REGION Network 10: Main Water Pump
   RUNG wire#powerrail
      #VFD_WaterPump(tInTimeout := t#5s, iInMode := #iInMode, iInAddress := 100, bInEstop := #bInEstop, bInSignalContactor := "I_WaterPumpContactorAux", bInEnableForward := #bWaterPumpInterlockOk, bInEnableReverse := false, rInCommandSpeed := 80.0, rInRampUpTime := 5.0, rInRampDownTime := 5.0, bInCommandForward := #bStartPumpCommand, bInCommandReverse := false, bInResetError := #bInResetError, bInMotorProtector := "I_WaterPumpMSP", bInLocalDisconnect := "I_WaterPumpDisconnect", bInClutch := true, bInCoolingFan := "I_WaterPumpCoolingFan", bInUseCurrentAlarm := true, bInUseMaxFrequencyAlarm := true, HMI_VFD_Control := "dbWaterSystem".VFD_WaterPump, rOutSpeed => #rPumpActualSpeed, rOutCurrent => #rPumpActualCurrent, rOutPower => #rPumpActualPower, bOutContactor => "Q_WaterPumpContactor", bOutForward => #bTemp, bOutReverse => #bTemp, bOutAuto => #bTemp, bOutError => #bTemp, ERROR_VFD => "dbErrors_WaterSystem".VFD_WaterPump)
   END_RUNG
   // the same network as SCL:
   #VFD_WaterPump(tInTimeout := t#5s,   // "fbVFD_GSeries"
                  iInMode := #iInMode,
                  iInAddress := 100,
                  bInEstop := #bInEstop,
                  bInSignalContactor := "I_WaterPumpContactorAux",
                  bInEnableForward := #bWaterPumpInterlockOk,
                  bInEnableReverse := false,
                  rInCommandSpeed := 80.0,
                  rInRampUpTime := 5.0,
                  rInRampDownTime := 5.0,
                  bInCommandForward := #bStartPumpCommand,
                  bInCommandReverse := false,
                  bInResetError := #bInResetError,
                  bInMotorProtector := "I_WaterPumpMSP",
                  bInLocalDisconnect := "I_WaterPumpDisconnect",
                  bInClutch := true,
                  bInCoolingFan := "I_WaterPumpCoolingFan",
                  bInUseCurrentAlarm := true,
                  bInUseMaxFrequencyAlarm := true,
                  HMI_VFD_Control := "dbWaterSystem".VFD_WaterPump,
                  rOutSpeed => #rPumpActualSpeed,
                  rOutCurrent => #rPumpActualCurrent,
                  rOutPower => #rPumpActualPower,
                  bOutContactor => "Q_WaterPumpContactor",
                  bOutForward => #bTemp,
                  bOutReverse => #bTemp,
                  bOutAuto => #bTemp,
                  bOutError => #bTemp,
                  ERROR_VFD => "dbErrors_WaterSystem".VFD_WaterPump);
END_REGION

REGION Network 11: Return Water Pump
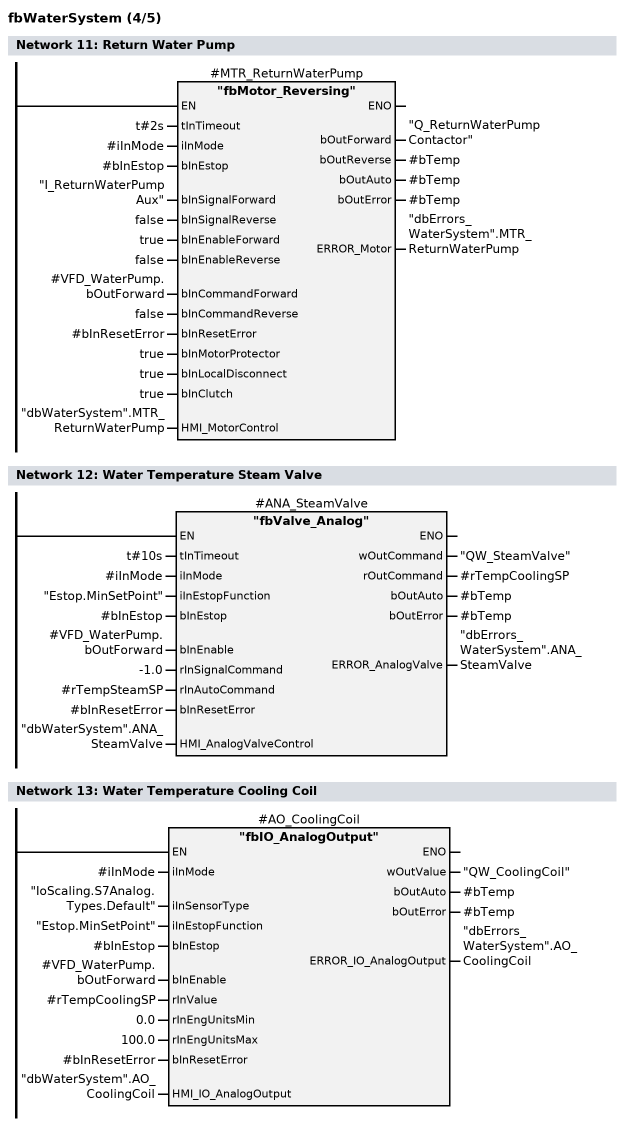
   RUNG wire#powerrail
      #MTR_ReturnWaterPump(tInTimeout := t#2s, iInMode := #iInMode, bInEstop := #bInEstop, bInSignalForward := "I_ReturnWaterPumpAux", bInSignalReverse := false, bInEnableForward := true, bInEnableReverse := false, bInCommandForward := #VFD_WaterPump.bOutForward, bInCommandReverse := false, bInResetError := #bInResetError, bInMotorProtector := true, bInLocalDisconnect := true, bInClutch := true, HMI_MotorControl := "dbWaterSystem".MTR_ReturnWaterPump, bOutForward => "Q_ReturnWaterPumpContactor", bOutReverse => #bTemp, bOutAuto => #bTemp, bOutError => #bTemp, ERROR_Motor => "dbErrors_WaterSystem".MTR_ReturnWaterPump)
   END_RUNG
   // the same network as SCL:
   #MTR_ReturnWaterPump(tInTimeout := t#2s,   // "fbMotor_Reversing"
                        iInMode := #iInMode,
                        bInEstop := #bInEstop,
                        bInSignalForward := "I_ReturnWaterPumpAux",
                        bInSignalReverse := false,
                        bInEnableForward := true,
                        bInEnableReverse := false,
                        bInCommandForward := #VFD_WaterPump.bOutForward,
                        bInCommandReverse := false,
                        bInResetError := #bInResetError,
                        bInMotorProtector := true,
                        bInLocalDisconnect := true,
                        bInClutch := true,
                        HMI_MotorControl := "dbWaterSystem".MTR_ReturnWaterPump,
                        bOutForward => "Q_ReturnWaterPumpContactor",
                        bOutReverse => #bTemp,
                        bOutAuto => #bTemp,
                        bOutError => #bTemp,
                        ERROR_Motor => "dbErrors_WaterSystem".MTR_ReturnWaterPump);
END_REGION

REGION Network 12: Water Temperature Steam Valve
   RUNG wire#powerrail
      #ANA_SteamValve(tInTimeout := t#10s, iInMode := #iInMode, iInEstopFunction := "Estop.MinSetPoint", bInEstop := #bInEstop, bInEnable := #VFD_WaterPump.bOutForward, rInSignalCommand := -1.0, rInAutoCommand := #rTempSteamSP, bInResetError := #bInResetError, HMI_AnalogValveControl := "dbWaterSystem".ANA_SteamValve, wOutCommand => "QW_SteamValve", rOutCommand => #rTempCoolingSP, bOutAuto => #bTemp, bOutError => #bTemp, ERROR_AnalogValve => "dbErrors_WaterSystem".ANA_SteamValve)
   END_RUNG
   // the same network as SCL:
   #ANA_SteamValve(tInTimeout := t#10s,   // "fbValve_Analog"
                   iInMode := #iInMode,
                   iInEstopFunction := "Estop.MinSetPoint",
                   bInEstop := #bInEstop,
                   bInEnable := #VFD_WaterPump.bOutForward,
                   rInSignalCommand := -1.0,
                   rInAutoCommand := #rTempSteamSP,
                   bInResetError := #bInResetError,
                   HMI_AnalogValveControl := "dbWaterSystem".ANA_SteamValve,
                   wOutCommand => "QW_SteamValve",
                   rOutCommand => #rTempCoolingSP,
                   bOutAuto => #bTemp,
                   bOutError => #bTemp,
                   ERROR_AnalogValve => "dbErrors_WaterSystem".ANA_SteamValve);
END_REGION

REGION Network 13: Water Temperature Cooling Coil
   RUNG wire#powerrail
      #AO_CoolingCoil(iInMode := #iInMode, iInSensorType := "IoScaling.S7Analog.Types.Default", iInEstopFunction := "Estop.MinSetPoint", bInEstop := #bInEstop, bInEnable := #VFD_WaterPump.bOutForward, rInValue := #rTempCoolingSP, rInEngUnitsMin := 0.0, rInEngUnitsMax := 100.0, bInResetError := #bInResetError, HMI_IO_AnalogOutput := "dbWaterSystem".AO_CoolingCoil, wOutValue => "QW_CoolingCoil", bOutAuto => #bTemp, bOutError => #bTemp, ERROR_IO_AnalogOutput => "dbErrors_WaterSystem".AO_CoolingCoil)
   END_RUNG
   // the same network as SCL:
   #AO_CoolingCoil(iInMode := #iInMode,   // "fbIO_AnalogOutput"
                   iInSensorType := "IoScaling.S7Analog.Types.Default",
                   iInEstopFunction := "Estop.MinSetPoint",
                   bInEstop := #bInEstop,
                   bInEnable := #VFD_WaterPump.bOutForward,
                   rInValue := #rTempCoolingSP,
                   rInEngUnitsMin := 0.0,
                   rInEngUnitsMax := 100.0,
                   bInResetError := #bInResetError,
                   HMI_IO_AnalogOutput := "dbWaterSystem".AO_CoolingCoil,
                   wOutValue => "QW_CoolingCoil",
                   bOutAuto => #bTemp,
                   bOutError => #bTemp,
                   ERROR_IO_AnalogOutput => "dbErrors_WaterSystem".AO_CoolingCoil);
END_REGION

REGION Network 14: -------------------------------------------------------- Alarms -----------------------------------------------------------------
END_REGION

REGION Network 15: Main Water Pump Pressure Alarm
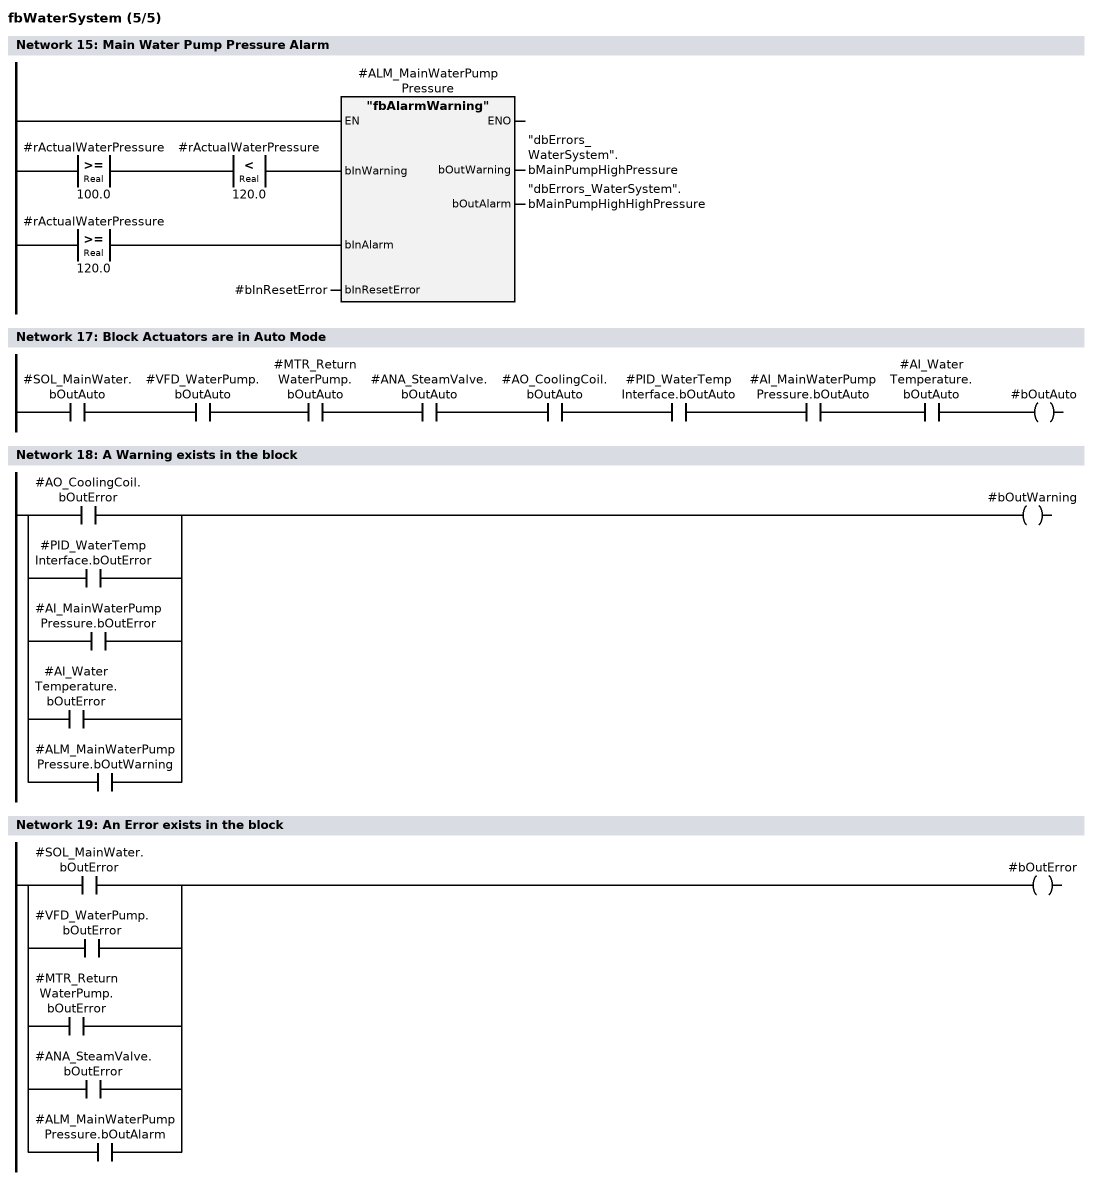
   RUNG wire#powerrail
      #ALM_MainWaterPumpPressure(bInWarning := wire#w1, bInAlarm := wire#w2, bInResetError := #bInResetError, bOutWarning => "dbErrors_WaterSystem".bMainPumpHighPressure, bOutAlarm => "dbErrors_WaterSystem".bMainPumpHighHighPressure)
   END_RUNG
   RUNG wire#powerrail
      { S7_Templates := "SrcType := Real" } GE_Contact(in1 := #rActualWaterPressure, in2 := 100.0)
      { S7_Templates := "SrcType := Real" } LT_Contact(in1 := #rActualWaterPressure, in2 := 120.0)
   END_RUNG wire#w1
   RUNG wire#powerrail
      { S7_Templates := "SrcType := Real" } GE_Contact(in1 := #rActualWaterPressure, in2 := 120.0)
   END_RUNG wire#w2
   // the same network as SCL:
   #ALM_MainWaterPumpPressure(bInWarning := (#rActualWaterPressure >= 100.0) AND (#rActualWaterPressure < 120.0),   // "fbAlarmWarning"
                           bInAlarm := #rActualWaterPressure >= 120.0,
                           bInResetError := #bInResetError,
                           bOutWarning => "dbErrors_WaterSystem".bMainPumpHighPressure,
                           bOutAlarm => "dbErrors_WaterSystem".bMainPumpHighHighPressure);
END_REGION

REGION Network 16: -------------------------------------------------------- Outputs -----------------------------------------------------------------
END_REGION

REGION Network 17: Block Actuators are in Auto Mode
   RUNG wire#powerrail
      Contact( #SOL_MainWater.bOutAuto )
      Contact( #VFD_WaterPump.bOutAuto )
      Contact( #MTR_ReturnWaterPump.bOutAuto )
      Contact( #ANA_SteamValve.bOutAuto )
      Contact( #AO_CoolingCoil.bOutAuto )
      Contact( #PID_WaterTempInterface.bOutAuto )
      Contact( #AI_MainWaterPumpPressure.bOutAuto )
      Contact( #AI_WaterTemperature.bOutAuto )
      Coil( #bOutAuto )
   END_RUNG
   // the same network as SCL:
   #bOutAuto := #SOL_MainWater.bOutAuto AND #VFD_WaterPump.bOutAuto AND #MTR_ReturnWaterPump.bOutAuto AND #ANA_SteamValve.bOutAuto AND #AO_CoolingCoil.bOutAuto AND #PID_WaterTempInterface.bOutAuto AND #AI_MainWaterPumpPressure.bOutAuto AND #AI_WaterTemperature.bOutAuto;
END_REGION

REGION Network 18: A Warning exists in the block
   RUNG wire#powerrail
      Contact( #AO_CoolingCoil.bOutError )
      wire#w1
      Coil( #bOutWarning )
   END_RUNG
   RUNG wire#powerrail
      Contact( #PID_WaterTempInterface.bOutError )
   END_RUNG wire#w1
   RUNG wire#powerrail
      Contact( #AI_MainWaterPumpPressure.bOutError )
   END_RUNG wire#w1
   RUNG wire#powerrail
      Contact( #AI_WaterTemperature.bOutError )
   END_RUNG wire#w1
   RUNG wire#powerrail
      Contact( #ALM_MainWaterPumpPressure.bOutWarning )
   END_RUNG wire#w1
   // the same network as SCL:
   #bOutWarning := #AO_CoolingCoil.bOutError OR #PID_WaterTempInterface.bOutError OR #AI_MainWaterPumpPressure.bOutError OR #AI_WaterTemperature.bOutError OR #ALM_MainWaterPumpPressure.bOutWarning;
END_REGION

REGION Network 19: An Error exists in the block
   RUNG wire#powerrail
      Contact( #SOL_MainWater.bOutError )
      wire#w1
      Coil( #bOutError )
   END_RUNG
   RUNG wire#powerrail
      Contact( #VFD_WaterPump.bOutError )
   END_RUNG wire#w1
   RUNG wire#powerrail
      Contact( #MTR_ReturnWaterPump.bOutError )
   END_RUNG wire#w1
   RUNG wire#powerrail
      Contact( #ANA_SteamValve.bOutError )
   END_RUNG wire#w1
   RUNG wire#powerrail
      Contact( #ALM_MainWaterPumpPressure.bOutAlarm )
   END_RUNG wire#w1
   // the same network as SCL:
   #bOutError := #SOL_MainWater.bOutError OR #VFD_WaterPump.bOutError OR #MTR_ReturnWaterPump.bOutError OR #ANA_SteamValve.bOutError OR #ALM_MainWaterPumpPressure.bOutAlarm;
END_REGION
END_FUNCTION_BLOCK

FUNCTION_BLOCK "fbAirSystem"   // FB520, LAD
TITLE = Air System Function Block
{ S7_Optimized_Access := 'FALSE' }
VERSION : 0.1
BEGIN

REGION Network 1: --------------------------------------------------------- Inputs ------------------------------------------------------------------
END_REGION

REGION Network 2: --------------------------------------------------- System Logic ------------------------------------------------------------
END_REGION

REGION Network 3: -------------------------------------------------------- Devices -----------------------------------------------------------------
END_REGION

REGION Network 4: Recirculation Fan
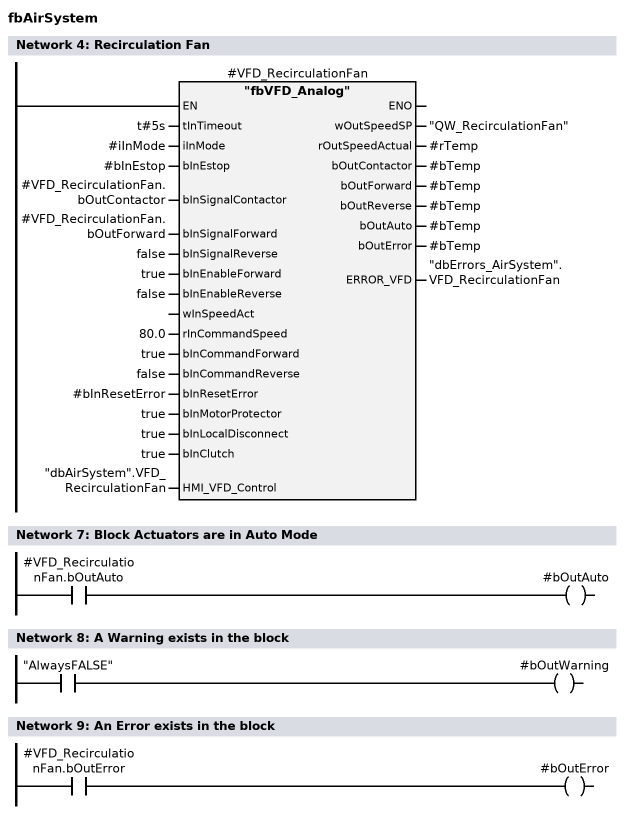
   RUNG wire#powerrail
      #VFD_RecirculationFan(tInTimeout := t#5s, iInMode := #iInMode, bInEstop := #bInEstop, bInSignalContactor := #VFD_RecirculationFan.bOutContactor, bInSignalForward := #VFD_RecirculationFan.bOutForward, bInSignalReverse := false, bInEnableForward := true, bInEnableReverse := false, wInSpeedAct :=, rInCommandSpeed := 80.0, bInCommandForward := true, bInCommandReverse := false, bInResetError := #bInResetError, bInMotorProtector := true, bInLocalDisconnect := true, bInClutch := true, HMI_VFD_Control := "dbAirSystem".VFD_RecirculationFan, wOutSpeedSP => "QW_RecirculationFan", rOutSpeedActual => #rTemp, bOutContactor => #bTemp, bOutForward => #bTemp, bOutReverse => #bTemp, bOutAuto => #bTemp, bOutError => #bTemp, ERROR_VFD => "dbErrors_AirSystem".VFD_RecirculationFan)
   END_RUNG
   // the same network as SCL:
   #VFD_RecirculationFan(tInTimeout := t#5s,   // "fbVFD_Analog"
                         iInMode := #iInMode,
                         bInEstop := #bInEstop,
                         bInSignalContactor := #VFD_RecirculationFan.bOutContactor,
                         bInSignalForward := #VFD_RecirculationFan.bOutForward,
                         bInSignalReverse := false,
                         bInEnableForward := true,
                         bInEnableReverse := false,
                         rInCommandSpeed := 80.0,
                         bInCommandForward := true,
                         bInCommandReverse := false,
                         bInResetError := #bInResetError,
                         bInMotorProtector := true,
                         bInLocalDisconnect := true,
                         bInClutch := true,
                         HMI_VFD_Control := "dbAirSystem".VFD_RecirculationFan,
                         wOutSpeedSP => "QW_RecirculationFan",
                         rOutSpeedActual => #rTemp,
                         bOutContactor => #bTemp,
                         bOutForward => #bTemp,
                         bOutReverse => #bTemp,
                         bOutAuto => #bTemp,
                         bOutError => #bTemp,
                         ERROR_VFD => "dbErrors_AirSystem".VFD_RecirculationFan);
END_REGION

REGION Network 5: -------------------------------------------------------- Alarms -----------------------------------------------------------------
END_REGION

REGION Network 6: -------------------------------------------------------- Outputs -----------------------------------------------------------------
END_REGION

REGION Network 7: Block Actuators are in Auto Mode
   RUNG wire#powerrail
      Contact( #VFD_RecirculationFan.bOutAuto )
      Coil( #bOutAuto )
   END_RUNG
   // the same network as SCL:
   #bOutAuto := #VFD_RecirculationFan.bOutAuto;
END_REGION

REGION Network 8: A Warning exists in the block
   RUNG wire#powerrail
      Contact( "AlwaysFALSE" )
      Coil( #bOutWarning )
   END_RUNG
   // the same network as SCL:
   #bOutWarning := "AlwaysFALSE";
END_REGION

REGION Network 9: An Error exists in the block
   RUNG wire#powerrail
      Contact( #VFD_RecirculationFan.bOutError )
      Coil( #bOutError )
   END_RUNG
   // the same network as SCL:
   #bOutError := #VFD_RecirculationFan.bOutError;
END_REGION
END_FUNCTION_BLOCK

// folder: Top Level

FUNCTION_BLOCK "fbCyclicInterrupt"   // FB30, LAD
TITLE = Cyclic Interrupt Function - 100ms
{ S7_Optimized_Access := 'FALSE' }
VERSION : 0.1
BEGIN

REGION Network 1: Call Temperature Control PID Block
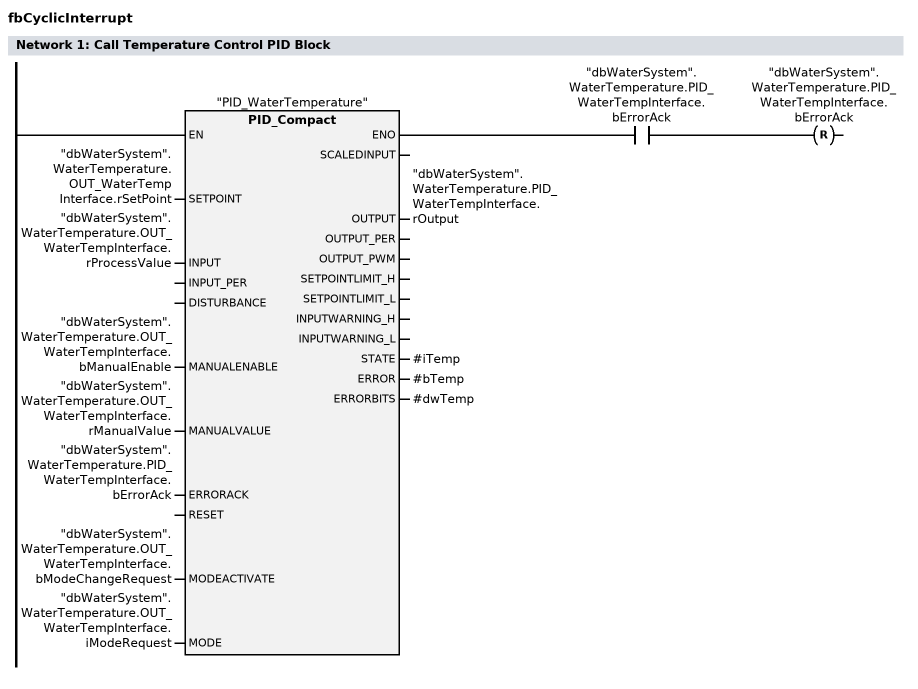
   // ENO of a box is taken as its EN; it also drops when the box reports an error
   "PID_WaterTemperature"(Setpoint := "dbWaterSystem".WaterTemperature.OUT_WaterTempInterface.rSetPoint,   // PID_Compact
                          Input := "dbWaterSystem".WaterTemperature.OUT_WaterTempInterface.rProcessValue,
                          ManualEnable := "dbWaterSystem".WaterTemperature.OUT_WaterTempInterface.bManualEnable,
                          ManualValue := "dbWaterSystem".WaterTemperature.OUT_WaterTempInterface.rManualValue,
                          ErrorAck := "dbWaterSystem".WaterTemperature.PID_WaterTempInterface.bErrorAck,
                          ModeActivate := "dbWaterSystem".WaterTemperature.OUT_WaterTempInterface.bModeChangeRequest,
                          Mode := "dbWaterSystem".WaterTemperature.OUT_WaterTempInterface.iModeRequest,
                          Output => "dbWaterSystem".WaterTemperature.PID_WaterTempInterface.rOutput,
                          State => #iTemp,
                          Error => #bTemp,
                          ErrorBits => #dwTemp);
   IF "dbWaterSystem".WaterTemperature.PID_WaterTempInterface.bErrorAck THEN
       "dbWaterSystem".WaterTemperature.PID_WaterTempInterface.bErrorAck := FALSE;
   END_IF;
END_REGION
END_FUNCTION_BLOCK

FUNCTION_BLOCK "fbMaster"   // FB500, LAD
TITLE = Master Function Block
{ S7_Optimized_Access := 'FALSE' }
VERSION : 0.1
   VAR_TEMP   // added for the SCL form of the ladder/FBD networks
      _w1 : Bool;
   END_VAR
BEGIN

REGION Network 1: Read HMI Push Buttons
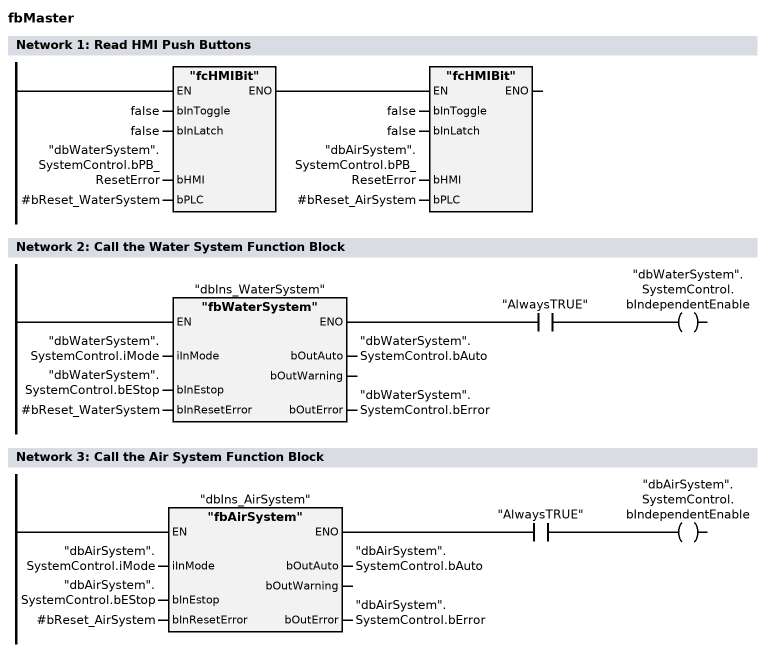
   RUNG wire#powerrail
      "fcHMIBit"(bInToggle := false, bInLatch := false, bHMI := "dbWaterSystem".SystemControl.bPB_ResetError, bPLC := #bReset_WaterSystem)
      "fcHMIBit"(bInToggle := false, bInLatch := false, bHMI := "dbAirSystem".SystemControl.bPB_ResetError, bPLC := #bReset_AirSystem)
   END_RUNG
   // the same network as SCL:
   "fcHMIBit"(bInToggle := false,
              bInLatch := false,
              bHMI := "dbWaterSystem".SystemControl.bPB_ResetError,
              bPLC := #bReset_WaterSystem,
              ENO => #_w1);
   IF #_w1 THEN
       "fcHMIBit"(bInToggle := false,
                  bInLatch := false,
                  bHMI := "dbAirSystem".SystemControl.bPB_ResetError,
                  bPLC := #bReset_AirSystem);
   END_IF;
END_REGION

REGION Network 2: Call the Water System Function Block
   RUNG wire#powerrail
      "dbIns_WaterSystem"(iInMode := "dbWaterSystem".SystemControl.iMode, bInEstop := "dbWaterSystem".SystemControl.bEStop, bInResetError := #bReset_WaterSystem, bOutAuto => "dbWaterSystem".SystemControl.bAuto, bOutWarning =>, bOutError => "dbWaterSystem".SystemControl.bError)
      Contact( "AlwaysTRUE" )
      Coil( "dbWaterSystem".SystemControl.bIndependentEnable )
   END_RUNG
   // the same network as SCL:
   "dbIns_WaterSystem"(iInMode := "dbWaterSystem".SystemControl.iMode,   // "fbWaterSystem"
                       bInEstop := "dbWaterSystem".SystemControl.bEStop,
                       bInResetError := #bReset_WaterSystem,
                       bOutAuto => "dbWaterSystem".SystemControl.bAuto,
                       bOutError => "dbWaterSystem".SystemControl.bError,
                       ENO => #_w1);
   "dbWaterSystem".SystemControl.bIndependentEnable := #_w1 AND "AlwaysTRUE";
END_REGION

REGION Network 3: Call the Air System Function Block
   RUNG wire#powerrail
      "dbIns_AirSystem"(iInMode := "dbAirSystem".SystemControl.iMode, bInEstop := "dbAirSystem".SystemControl.bEStop, bInResetError := #bReset_AirSystem, bOutAuto => "dbAirSystem".SystemControl.bAuto, bOutWarning =>, bOutError => "dbAirSystem".SystemControl.bError)
      Contact( "AlwaysTRUE" )
      Coil( "dbAirSystem".SystemControl.bIndependentEnable )
   END_RUNG
   // the same network as SCL:
   "dbIns_AirSystem"(iInMode := "dbAirSystem".SystemControl.iMode,   // "fbAirSystem"
                     bInEstop := "dbAirSystem".SystemControl.bEStop,
                     bInResetError := #bReset_AirSystem,
                     bOutAuto => "dbAirSystem".SystemControl.bAuto,
                     bOutError => "dbAirSystem".SystemControl.bError,
                     ENO => #_w1);
   "dbAirSystem".SystemControl.bIndependentEnable := #_w1 AND "AlwaysTRUE";
END_REGION
END_FUNCTION_BLOCK

// ===== library types =====

// folder: Resources/Conversion

FUNCTION "fcByteToBits" : Void   // FC302, SCL
TITLE = Decode byte
{ S7_Optimized_Access := 'FALSE' }
AUTHOR : Boris
VERSION : 1.0
BEGIN

   #TEMPBYTE    := #byInByte;
   #bOutBit00  := #TEMPARRAY[0];
   #bOutBit01  := #TEMPARRAY[1];
   #bOutBit02  := #TEMPARRAY[2];
   #bOutBit03  := #TEMPARRAY[3];
   #bOutBit04  := #TEMPARRAY[4];
   #bOutBit05  := #TEMPARRAY[5];
   #bOutBit06  := #TEMPARRAY[6];
   #bOutBit07  := #TEMPARRAY[7];

   ENO := true;
END_FUNCTION

FUNCTION "fcBitsToByte" : Void   // FC303, SCL
TITLE = Pack Bits into byte
{ S7_Optimized_Access := 'FALSE' }
AUTHOR : Boris
VERSION : 1.0
BEGIN

       #TEMPARRAY[0] := #bInBit00;
       #TEMPARRAY[1] := #bInBit01;
       #TEMPARRAY[2] := #bInBit02;
       #TEMPARRAY[3] := #bInBit03;
       #TEMPARRAY[4] := #bInBit04;
       #TEMPARRAY[5] := #bInBit05;
       #TEMPARRAY[6] := #bInBit06;
       #TEMPARRAY[7] := #bInBit07;
       #byOutByte := #TEMPBYTE;

   ENO := true;
END_FUNCTION

FUNCTION "fcSwapWords" : Void   // FC303, LAD
TITLE = Swaps the words in a DWORD
{ S7_Optimized_Access := 'FALSE' }
AUTHOR : DMC
FAMILY : LowLevel
VERSION : 0.1
BEGIN

REGION Network 1: Swap the Words
   // High word and Low word are swapped
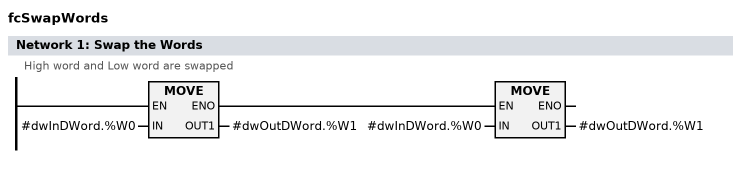
   RUNG wire#powerrail
      { S7_GenerateENO := "TRUE" } Move(in := #dwInDWord.%W0, out1 => #dwOutDWord.%W1)
      { S7_GenerateENO := "TRUE" } Move(in := #dwInDWord.%W0, out1 => #dwOutDWord.%W1)
   END_RUNG
   // the same network as SCL:
   // ENO of a box is taken as its EN; it also drops when the box reports an error
   #dwOutDWord.%W1 := #dwInDWord.%W0;
   #dwOutDWord.%W1 := #dwInDWord.%W0;
END_REGION
END_FUNCTION

FUNCTION "fcSwapWords" : Void   // FC307, SCL
{ S7_Optimized_Access := 'FALSE' }
VERSION : 0.1
BEGIN
   #TEMPDWORDIN := #dwInDWord;
   #TEMPARRAYOUT[0] := #TEMPARRAYIN[1];
   #TEMPARRAYOUT[1] := #TEMPARRAYIN[0];
   #dwOutDWord := #TEMPDWORDOUT;

   ENO := TRUE;
END_FUNCTION

FUNCTION "fcReal2Time_Min" : Void   // FC320, LAD
TITLE = Convert real value (minutes) to S7 Time
{ S7_Optimized_Access := 'FALSE' }
AUTHOR : DMC
FAMILY : LowLevel
VERSION : 0.1
BEGIN

REGION Network 1: Set Default time value to Zero
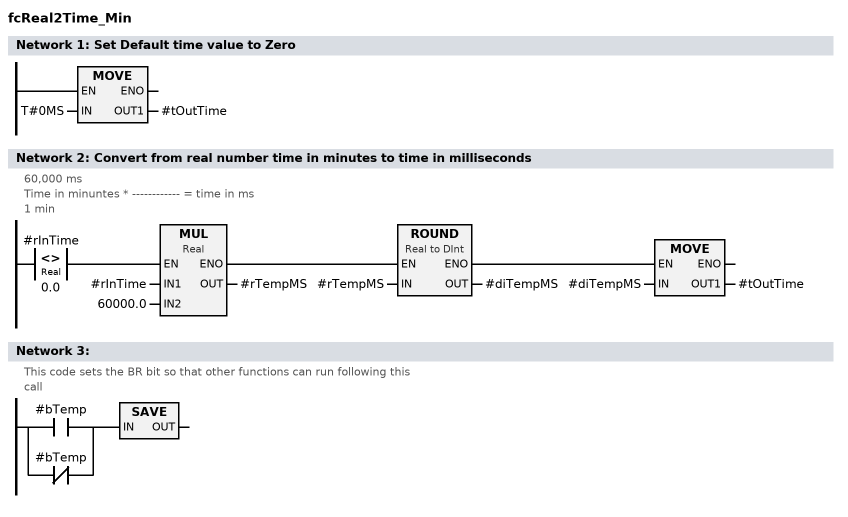
   RUNG wire#powerrail
      { S7_GenerateENO := "TRUE" } Move(in := T#0MS, out1 => #tOutTime)
   END_RUNG
   // the same network as SCL:
   #tOutTime := T#0MS;
END_REGION

REGION Network 2: Convert from real number time in minutes to time in milliseconds
   // 60,000 ms
   // Time in minuntes * ------------ = time in ms
   //                       1 min
   RUNG wire#powerrail
      { S7_Templates := "SrcType := Real" } NE_Contact(in1 := #rInTime, in2 := 0.0)
      { S7_Templates := "SrcType := Real"; S7_GenerateENO := "TRUE" } Mul(in1 := #rInTime, in2 := 60000.0, out => #rTempMS)
      { S7_Templates := "[SrcType := Real, DestType := DInt]"; S7_GenerateENO := "TRUE" } Round(in := #rTempMS, out => #diTempMS)
      { S7_GenerateENO := "TRUE" } Move(in := #diTempMS, out1 => #tOutTime)
   END_RUNG
   // the same network as SCL:
   // ENO of a box is taken as its EN; it also drops when the box reports an error
   IF #rInTime <> 0.0 THEN
       #rTempMS := #rInTime * 60000.0;
       #diTempMS := ROUND(#rTempMS);
       #tOutTime := #diTempMS;
   END_IF;
END_REGION

REGION Network 3
   // This code sets the BR bit so that other functions can run following this 
   // call
   // no SCL statement known for Save: written as a call
   Save(in := #bTemp OR NOT #bTemp);
END_REGION
END_FUNCTION

FUNCTION "fcReal2Time_Min" : Void   // FC320, LAD
TITLE = Convert real value (minutes) to S7 Time
{ S7_Optimized_Access := 'FALSE' }
AUTHOR : DMC
FAMILY : LowLevel
VERSION : 0.1
BEGIN

REGION Network 1: Set Default time value to Zero
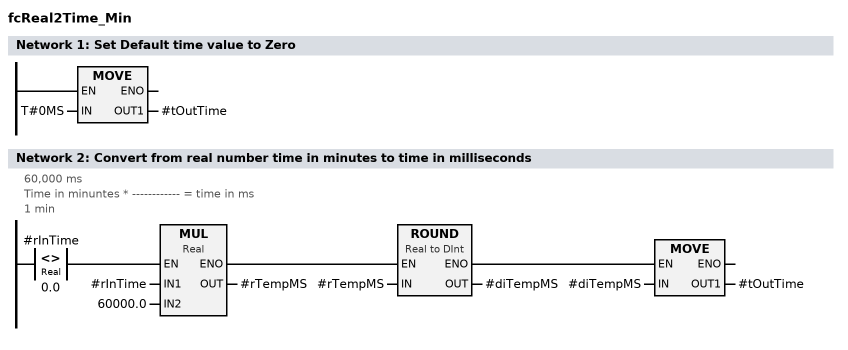
   RUNG wire#powerrail
      { S7_GenerateENO := "TRUE" } Move(in := T#0MS, out1 => #tOutTime)
   END_RUNG
   // the same network as SCL:
   #tOutTime := T#0MS;
END_REGION

REGION Network 2: Convert from real number time in minutes to time in milliseconds
   // 60,000 ms
   // Time in minuntes * ------------ = time in ms
   //                       1 min
   RUNG wire#powerrail
      { S7_Templates := "SrcType := Real" } NE_Contact(in1 := #rInTime, in2 := 0.0)
      { S7_Templates := "SrcType := Real"; S7_GenerateENO := "TRUE" } Mul(in1 := #rInTime, in2 := 60000.0, out => #rTempMS)
      { S7_Templates := "[SrcType := Real, DestType := DInt]"; S7_GenerateENO := "TRUE" } Round(in := #rTempMS, out => #diTempMS)
      { S7_GenerateENO := "TRUE" } Move(in := #diTempMS, out1 => #tOutTime)
   END_RUNG
   // the same network as SCL:
   // ENO of a box is taken as its EN; it also drops when the box reports an error
   IF #rInTime <> 0.0 THEN
       #rTempMS := #rInTime * 60000.0;
       #diTempMS := ROUND(#rTempMS);
       #tOutTime := #diTempMS;
   END_IF;
END_REGION
END_FUNCTION

FUNCTION "fcTime2Real_Min" : Void   // FC321, LAD
TITLE = Convert S7 time to real value (minutes)
{ S7_Optimized_Access := 'FALSE' }
AUTHOR : DMC
FAMILY : LowLevel
VERSION : 0.1
BEGIN

REGION Network 1: Load the time value and convert to a real
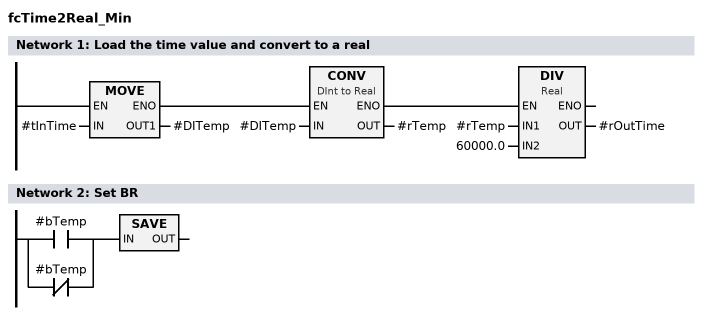
   RUNG wire#powerrail
      { S7_GenerateENO := "TRUE" } Move(in := #tInTime, out1 => #DITemp)
      { S7_Templates := "[SrcType := DInt, DestType := Real]"; S7_GenerateENO := "TRUE" } Convert(in := #DITemp, out => #rTemp)
      { S7_Templates := "SrcType := Real"; S7_GenerateENO := "TRUE" } Div(in1 := #rTemp, in2 := 60000.0, out => #rOutTime)
   END_RUNG
   // the same network as SCL:
   // ENO of a box is taken as its EN; it also drops when the box reports an error
   #DITemp := #tInTime;
   #rTemp := DINT_TO_REAL(#DITemp);
   #rOutTime := #rTemp / 60000.0;
END_REGION

REGION Network 2: Set BR
   // no SCL statement known for Save: written as a call
   Save(in := #bTemp OR NOT #bTemp);
END_REGION
END_FUNCTION

FUNCTION "fcTime2Real_Min" : Void   // FC321, LAD
TITLE = Convert S7 time to real value (minutes)
{ S7_Optimized_Access := 'FALSE' }
AUTHOR : DMC
FAMILY : LowLevel
VERSION : 0.1
BEGIN

REGION Network 1: Load the time value and convert to a real
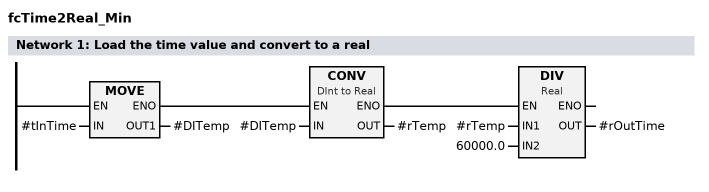
   RUNG wire#powerrail
      { S7_GenerateENO := "TRUE" } Move(in := #tInTime, out1 => #DITemp)
      { S7_Templates := "[SrcType := DInt, DestType := Real]"; S7_GenerateENO := "TRUE" } Convert(in := #DITemp, out => #rTemp)
      { S7_Templates := "SrcType := Real"; S7_GenerateENO := "TRUE" } Div(in1 := #rTemp, in2 := 60000.0, out => #rOutTime)
   END_RUNG
   // the same network as SCL:
   // ENO of a box is taken as its EN; it also drops when the box reports an error
   #DITemp := #tInTime;
   #rTemp := DINT_TO_REAL(#DITemp);
   #rOutTime := #rTemp / 60000.0;
END_REGION
END_FUNCTION

FUNCTION "fcReal2Time_Sec" : Void   // FC322, LAD
TITLE = Convert real value (minutes) to S7 Time
{ S7_Optimized_Access := 'FALSE' }
AUTHOR : DMC
FAMILY : LowLevel
VERSION : 0.1
BEGIN

REGION Network 1: Set Default time value to Zero
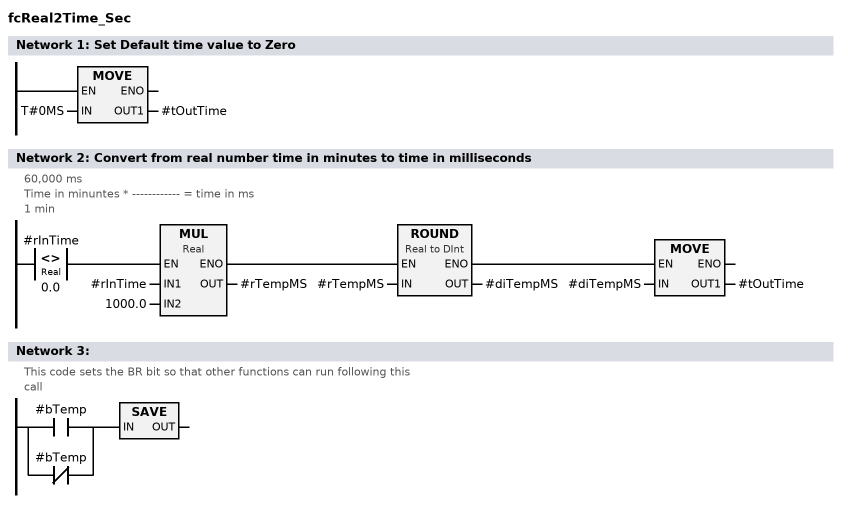
   RUNG wire#powerrail
      { S7_GenerateENO := "TRUE" } Move(in := T#0MS, out1 => #tOutTime)
   END_RUNG
   // the same network as SCL:
   #tOutTime := T#0MS;
END_REGION

REGION Network 2: Convert from real number time in minutes to time in milliseconds
   // 60,000 ms
   // Time in minuntes * ------------ = time in ms
   //                       1 min
   RUNG wire#powerrail
      { S7_Templates := "SrcType := Real" } NE_Contact(in1 := #rInTime, in2 := 0.0)
      { S7_Templates := "SrcType := Real"; S7_GenerateENO := "TRUE" } Mul(in1 := #rInTime, in2 := 1000.0, out => #rTempMS)
      { S7_Templates := "[SrcType := Real, DestType := DInt]"; S7_GenerateENO := "TRUE" } Round(in := #rTempMS, out => #diTempMS)
      { S7_GenerateENO := "TRUE" } Move(in := #diTempMS, out1 => #tOutTime)
   END_RUNG
   // the same network as SCL:
   // ENO of a box is taken as its EN; it also drops when the box reports an error
   IF #rInTime <> 0.0 THEN
       #rTempMS := #rInTime * 1000.0;
       #diTempMS := ROUND(#rTempMS);
       #tOutTime := #diTempMS;
   END_IF;
END_REGION

REGION Network 3
   // This code sets the BR bit so that other functions can run following this 
   // call
   // no SCL statement known for Save: written as a call
   Save(in := #bTemp OR NOT #bTemp);
END_REGION
END_FUNCTION

FUNCTION "fcReal2Time_Sec" : Void   // FC322, LAD
TITLE = Convert real value (minutes) to S7 Time
{ S7_Optimized_Access := 'FALSE' }
AUTHOR : DMC
FAMILY : LowLevel
VERSION : 0.1
BEGIN

REGION Network 1: Set Default time value to Zero
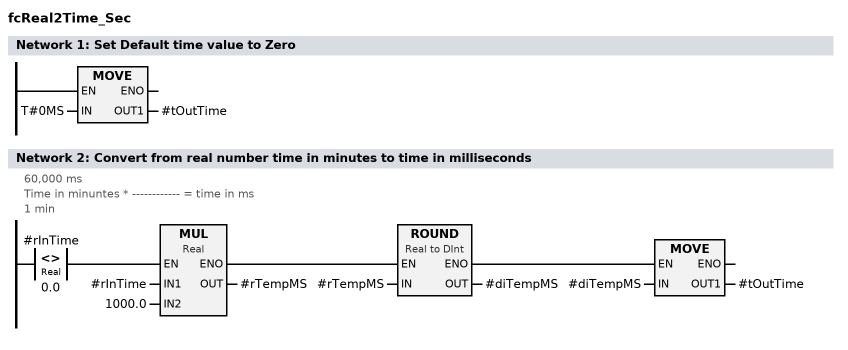
   RUNG wire#powerrail
      { S7_GenerateENO := "TRUE" } Move(in := T#0MS, out1 => #tOutTime)
   END_RUNG
   // the same network as SCL:
   #tOutTime := T#0MS;
END_REGION

REGION Network 2: Convert from real number time in minutes to time in milliseconds
   // 60,000 ms
   // Time in minuntes * ------------ = time in ms
   //                       1 min
   RUNG wire#powerrail
      { S7_Templates := "SrcType := Real" } NE_Contact(in1 := #rInTime, in2 := 0.0)
      { S7_Templates := "SrcType := Real"; S7_GenerateENO := "TRUE" } Mul(in1 := #rInTime, in2 := 1000.0, out => #rTempMS)
      { S7_Templates := "[SrcType := Real, DestType := DInt]"; S7_GenerateENO := "TRUE" } Round(in := #rTempMS, out => #diTempMS)
      { S7_GenerateENO := "TRUE" } Move(in := #diTempMS, out1 => #tOutTime)
   END_RUNG
   // the same network as SCL:
   // ENO of a box is taken as its EN; it also drops when the box reports an error
   IF #rInTime <> 0.0 THEN
       #rTempMS := #rInTime * 1000.0;
       #diTempMS := ROUND(#rTempMS);
       #tOutTime := #diTempMS;
   END_IF;
END_REGION
END_FUNCTION

FUNCTION "fcTime2Real_Sec" : Void   // FC323, LAD
TITLE = Convert S7 time to real value (minutes)
{ S7_Optimized_Access := 'FALSE' }
AUTHOR : DMC
FAMILY : LowLevel
VERSION : 0.1
BEGIN

REGION Network 1: Load the time value and convert to a real
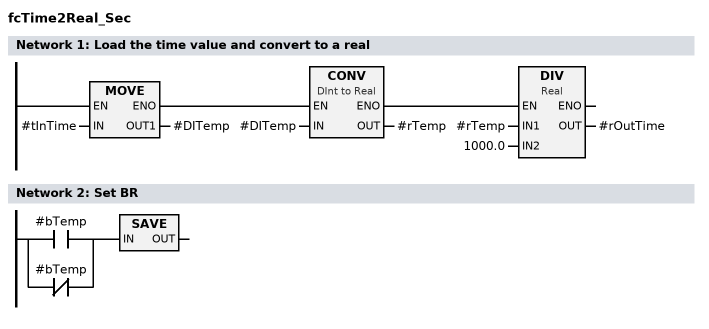
   RUNG wire#powerrail
      { S7_GenerateENO := "TRUE" } Move(in := #tInTime, out1 => #DITemp)
      { S7_Templates := "[SrcType := DInt, DestType := Real]"; S7_GenerateENO := "TRUE" } Convert(in := #DITemp, out => #rTemp)
      { S7_Templates := "SrcType := Real"; S7_GenerateENO := "TRUE" } Div(in1 := #rTemp, in2 := 1000.0, out => #rOutTime)
   END_RUNG
   // the same network as SCL:
   // ENO of a box is taken as its EN; it also drops when the box reports an error
   #DITemp := #tInTime;
   #rTemp := DINT_TO_REAL(#DITemp);
   #rOutTime := #rTemp / 1000.0;
END_REGION

REGION Network 2: Set BR
   // no SCL statement known for Save: written as a call
   Save(in := #bTemp OR NOT #bTemp);
END_REGION
END_FUNCTION

FUNCTION "fcTime2Real_Sec" : Void   // FC323, LAD
TITLE = Convert S7 time to real value (minutes)
{ S7_Optimized_Access := 'FALSE' }
AUTHOR : DMC
FAMILY : LowLevel
VERSION : 0.1
BEGIN

REGION Network 1: Load the time value and convert to a real
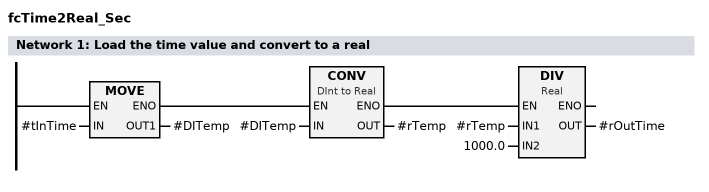
   RUNG wire#powerrail
      { S7_GenerateENO := "TRUE" } Move(in := #tInTime, out1 => #DITemp)
      { S7_Templates := "[SrcType := DInt, DestType := Real]"; S7_GenerateENO := "TRUE" } Convert(in := #DITemp, out => #rTemp)
      { S7_Templates := "SrcType := Real"; S7_GenerateENO := "TRUE" } Div(in1 := #rTemp, in2 := 1000.0, out => #rOutTime)
   END_RUNG
   // the same network as SCL:
   // ENO of a box is taken as its EN; it also drops when the box reports an error
   #DITemp := #tInTime;
   #rTemp := DINT_TO_REAL(#DITemp);
   #rOutTime := #rTemp / 1000.0;
END_REGION
END_FUNCTION

FUNCTION "fcTimeSplit" : Void   // FC326, LAD
TITLE = Parse Time Variable
{ S7_Optimized_Access := 'FALSE' }
VERSION : 0.1
BEGIN

REGION Network 1: Convert time to double int
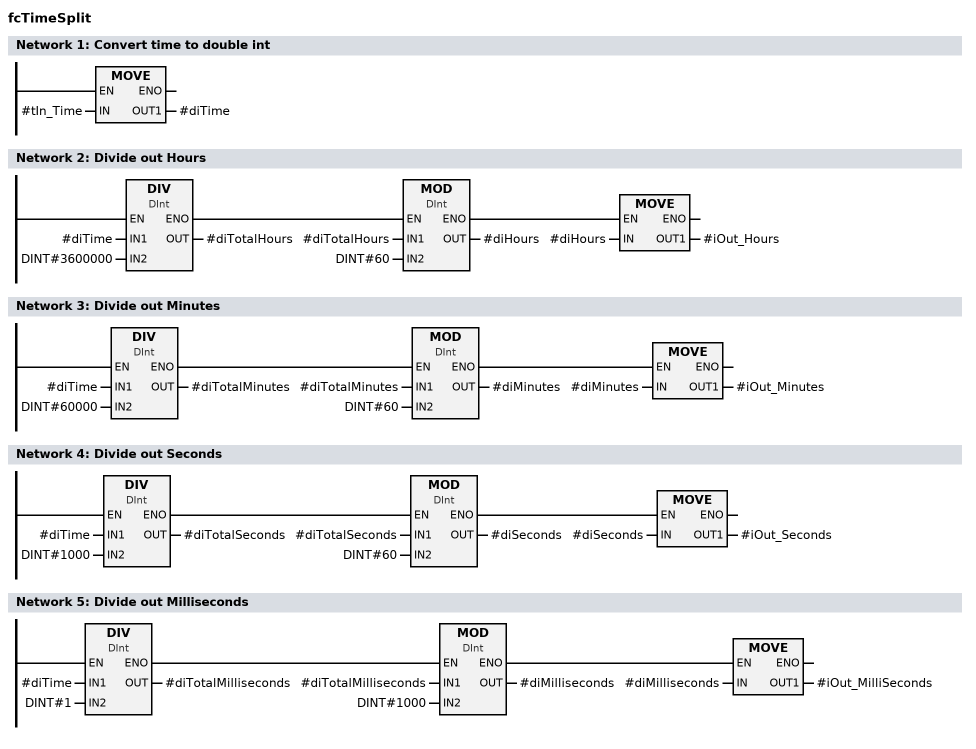
   RUNG wire#powerrail
      { S7_GenerateENO := "TRUE" } Move(in := #tIn_Time, out1 => #diTime)
   END_RUNG
   // the same network as SCL:
   #diTime := #tIn_Time;
END_REGION

REGION Network 2: Divide out Hours
   RUNG wire#powerrail
      { S7_Templates := "SrcType := DInt"; S7_GenerateENO := "TRUE" } Div(in1 := #diTime, in2 := DINT#3600000, out => #diTotalHours)
      { S7_Templates := "SrcType := DInt"; S7_GenerateENO := "TRUE" } Mod(in1 := #diTotalHours, in2 := DINT#60, out => #diHours)
      { S7_GenerateENO := "TRUE" } Move(in := #diHours, out1 => #iOut_Hours)
   END_RUNG
   // the same network as SCL:
   // ENO of a box is taken as its EN; it also drops when the box reports an error
   #diTotalHours := #diTime / DINT#3600000;
   #diHours := #diTotalHours MOD DINT#60;
   #iOut_Hours := #diHours;
END_REGION

REGION Network 3: Divide out Minutes
   RUNG wire#powerrail
      { S7_Templates := "SrcType := DInt"; S7_GenerateENO := "TRUE" } Div(in1 := #diTime, in2 := DINT#60000, out => #diTotalMinutes)
      { S7_Templates := "SrcType := DInt"; S7_GenerateENO := "TRUE" } Mod(in1 := #diTotalMinutes, in2 := DINT#60, out => #diMinutes)
      { S7_GenerateENO := "TRUE" } Move(in := #diMinutes, out1 => #iOut_Minutes)
   END_RUNG
   // the same network as SCL:
   // ENO of a box is taken as its EN; it also drops when the box reports an error
   #diTotalMinutes := #diTime / DINT#60000;
   #diMinutes := #diTotalMinutes MOD DINT#60;
   #iOut_Minutes := #diMinutes;
END_REGION

REGION Network 4: Divide out Seconds
   RUNG wire#powerrail
      { S7_Templates := "SrcType := DInt"; S7_GenerateENO := "TRUE" } Div(in1 := #diTime, in2 := DINT#1000, out => #diTotalSeconds)
      { S7_Templates := "SrcType := DInt"; S7_GenerateENO := "TRUE" } Mod(in1 := #diTotalSeconds, in2 := DINT#60, out => #diSeconds)
      { S7_GenerateENO := "TRUE" } Move(in := #diSeconds, out1 => #iOut_Seconds)
   END_RUNG
   // the same network as SCL:
   // ENO of a box is taken as its EN; it also drops when the box reports an error
   #diTotalSeconds := #diTime / DINT#1000;
   #diSeconds := #diTotalSeconds MOD DINT#60;
   #iOut_Seconds := #diSeconds;
END_REGION

REGION Network 5: Divide out Milliseconds
   RUNG wire#powerrail
      { S7_Templates := "SrcType := DInt"; S7_GenerateENO := "TRUE" } Div(in1 := #diTime, in2 := DINT#1, out => #diTotalMilliseconds)
      { S7_Templates := "SrcType := DInt"; S7_GenerateENO := "TRUE" } Mod(in1 := #diTotalMilliseconds, in2 := DINT#1000, out => #diMilliseconds)
      { S7_GenerateENO := "TRUE" } Move(in := #diMilliseconds, out1 => #iOut_MilliSeconds)
   END_RUNG
   // the same network as SCL:
   // ENO of a box is taken as its EN; it also drops when the box reports an error
   #diTotalMilliseconds := #diTime / DINT#1;
   #diMilliseconds := #diTotalMilliseconds MOD DINT#1000;
   #iOut_MilliSeconds := #diMilliseconds;
END_REGION
END_FUNCTION

FUNCTION "fcRead_Clk_Parts" : Void   // FC327, LAD
TITLE = Parse Date and Time Variable
{ S7_Optimized_Access := 'FALSE' }
VERSION : 0.1
BEGIN

REGION Network 1: Read Clock
